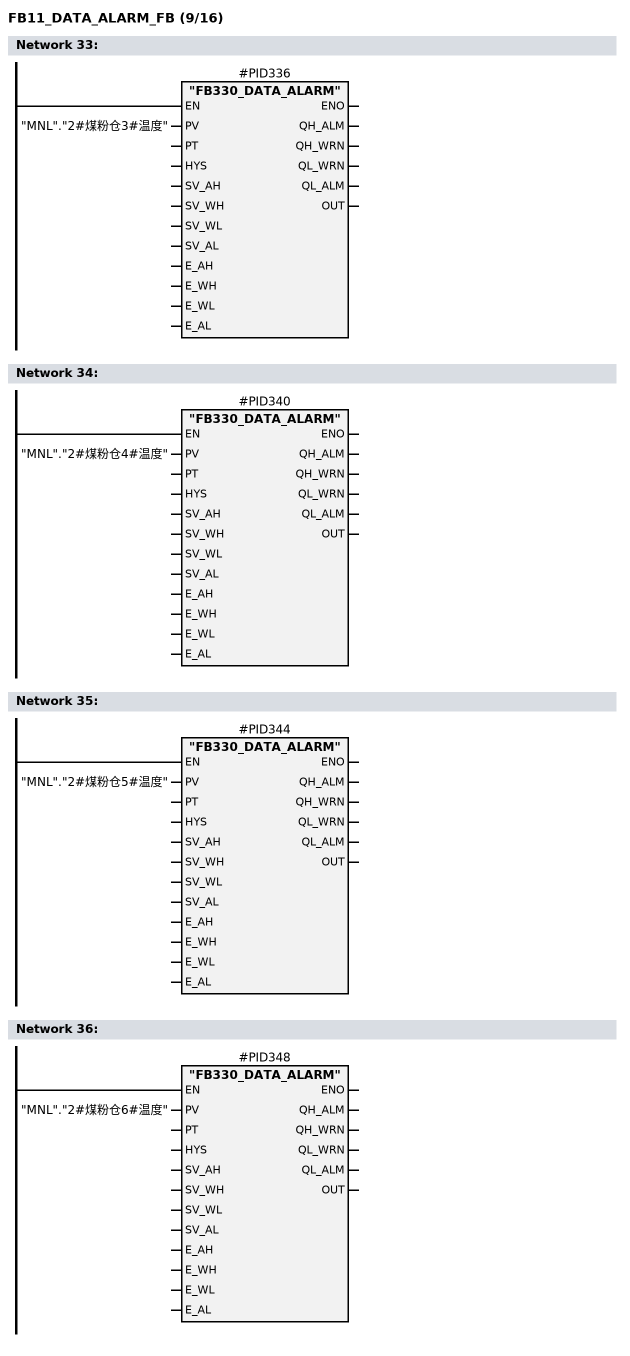
   RUNG wire#powerrail
      #PID336(PV := "MNL"."2#煤粉仓3#温度", PT :=, HYS :=, SV_AH :=, SV_WH :=, SV_WL :=, SV_AL :=, E_AH :=, E_WH :=, E_WL :=, E_AL :=, QH_ALM =>, QH_WRN =>, QL_WRN =>, QL_ALM =>, OUT =>)
   END_RUNG
   // the same network as SCL:
   #PID336(PV := "MNL"."2#煤粉仓3#温度");   // "FB330_DATA_ALARM"
END_REGION

REGION Network 34
   RUNG wire#powerrail
      #PID340(PV := "MNL"."2#煤粉仓4#温度", PT :=, HYS :=, SV_AH :=, SV_WH :=, SV_WL :=, SV_AL :=, E_AH :=, E_WH :=, E_WL :=, E_AL :=, QH_ALM =>, QH_WRN =>, QL_WRN =>, QL_ALM =>, OUT =>)
   END_RUNG
   // the same network as SCL:
   #PID340(PV := "MNL"."2#煤粉仓4#温度");   // "FB330_DATA_ALARM"
END_REGION

REGION Network 35
   RUNG wire#powerrail
      #PID344(PV := "MNL"."2#煤粉仓5#温度", PT :=, HYS :=, SV_AH :=, SV_WH :=, SV_WL :=, SV_AL :=, E_AH :=, E_WH :=, E_WL :=, E_AL :=, QH_ALM =>, QH_WRN =>, QL_WRN =>, QL_ALM =>, OUT =>)
   END_RUNG
   // the same network as SCL:
   #PID344(PV := "MNL"."2#煤粉仓5#温度");   // "FB330_DATA_ALARM"
END_REGION

REGION Network 36
   RUNG wire#powerrail
      #PID348(PV := "MNL"."2#煤粉仓6#温度", PT :=, HYS :=, SV_AH :=, SV_WH :=, SV_WL :=, SV_AL :=, E_AH :=, E_WH :=, E_WL :=, E_AL :=, QH_ALM =>, QH_WRN =>, QL_WRN =>, QL_ALM =>, OUT =>)
   END_RUNG
   // the same network as SCL:
   #PID348(PV := "MNL"."2#煤粉仓6#温度");   // "FB330_DATA_ALARM"
END_REGION

REGION Network 37
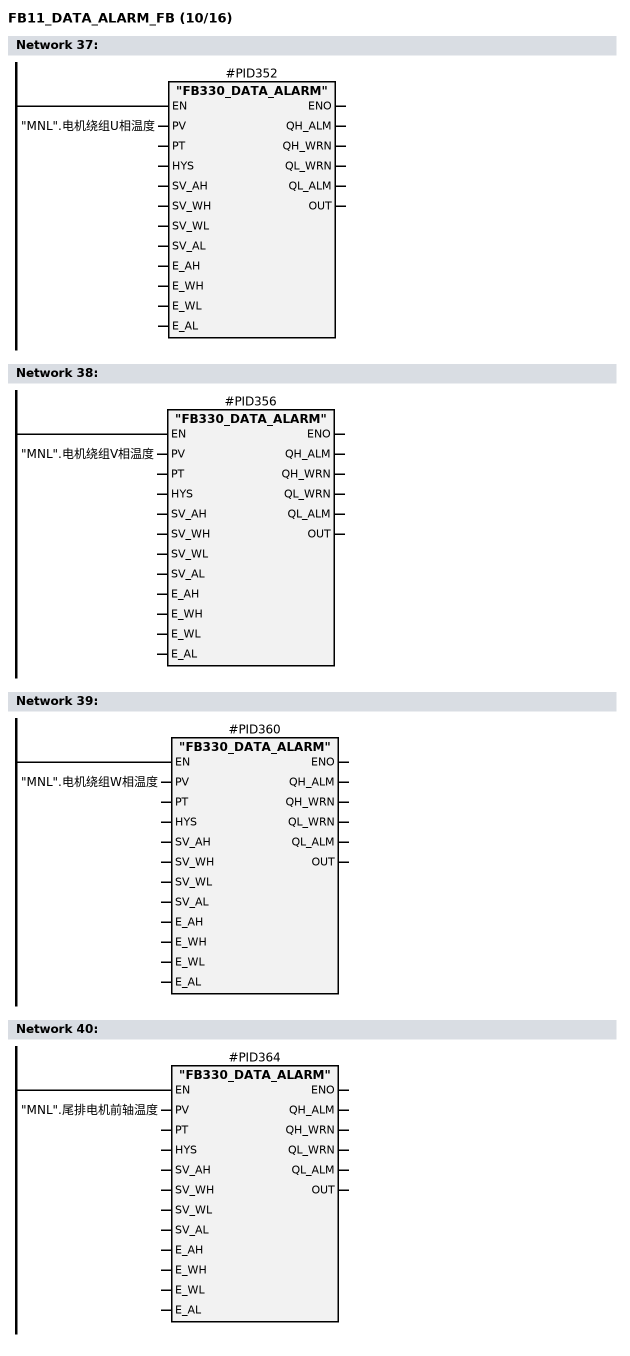
   RUNG wire#powerrail
      #PID352(PV := "MNL".电机绕组U相温度, PT :=, HYS :=, SV_AH :=, SV_WH :=, SV_WL :=, SV_AL :=, E_AH :=, E_WH :=, E_WL :=, E_AL :=, QH_ALM =>, QH_WRN =>, QL_WRN =>, QL_ALM =>, OUT =>)
   END_RUNG
   // the same network as SCL:
   #PID352(PV := "MNL".电机绕组U相温度);   // "FB330_DATA_ALARM"
END_REGION

REGION Network 38
   RUNG wire#powerrail
      #PID356(PV := "MNL".电机绕组V相温度, PT :=, HYS :=, SV_AH :=, SV_WH :=, SV_WL :=, SV_AL :=, E_AH :=, E_WH :=, E_WL :=, E_AL :=, QH_ALM =>, QH_WRN =>, QL_WRN =>, QL_ALM =>, OUT =>)
   END_RUNG
   // the same network as SCL:
   #PID356(PV := "MNL".电机绕组V相温度);   // "FB330_DATA_ALARM"
END_REGION

REGION Network 39
   RUNG wire#powerrail
      #PID360(PV := "MNL".电机绕组W相温度, PT :=, HYS :=, SV_AH :=, SV_WH :=, SV_WL :=, SV_AL :=, E_AH :=, E_WH :=, E_WL :=, E_AL :=, QH_ALM =>, QH_WRN =>, QL_WRN =>, QL_ALM =>, OUT =>)
   END_RUNG
   // the same network as SCL:
   #PID360(PV := "MNL".电机绕组W相温度);   // "FB330_DATA_ALARM"
END_REGION

REGION Network 40
   RUNG wire#powerrail
      #PID364(PV := "MNL".尾排电机前轴温度, PT :=, HYS :=, SV_AH :=, SV_WH :=, SV_WL :=, SV_AL :=, E_AH :=, E_WH :=, E_WL :=, E_AL :=, QH_ALM =>, QH_WRN =>, QL_WRN =>, QL_ALM =>, OUT =>)
   END_RUNG
   // the same network as SCL:
   #PID364(PV := "MNL".尾排电机前轴温度);   // "FB330_DATA_ALARM"
END_REGION

REGION Network 41
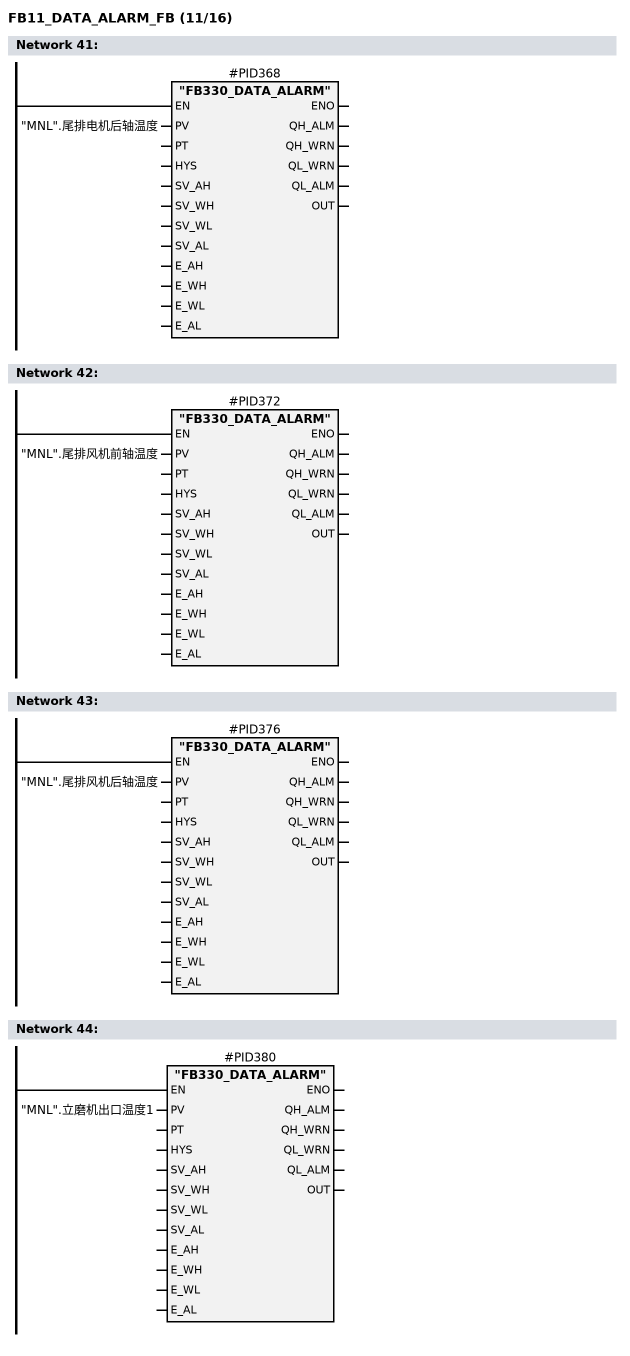
   RUNG wire#powerrail
      #PID368(PV := "MNL".尾排电机后轴温度, PT :=, HYS :=, SV_AH :=, SV_WH :=, SV_WL :=, SV_AL :=, E_AH :=, E_WH :=, E_WL :=, E_AL :=, QH_ALM =>, QH_WRN =>, QL_WRN =>, QL_ALM =>, OUT =>)
   END_RUNG
   // the same network as SCL:
   #PID368(PV := "MNL".尾排电机后轴温度);   // "FB330_DATA_ALARM"
END_REGION

REGION Network 42
   RUNG wire#powerrail
      #PID372(PV := "MNL".尾排风机前轴温度, PT :=, HYS :=, SV_AH :=, SV_WH :=, SV_WL :=, SV_AL :=, E_AH :=, E_WH :=, E_WL :=, E_AL :=, QH_ALM =>, QH_WRN =>, QL_WRN =>, QL_ALM =>, OUT =>)
   END_RUNG
   // the same network as SCL:
   #PID372(PV := "MNL".尾排风机前轴温度);   // "FB330_DATA_ALARM"
END_REGION

REGION Network 43
   RUNG wire#powerrail
      #PID376(PV := "MNL".尾排风机后轴温度, PT :=, HYS :=, SV_AH :=, SV_WH :=, SV_WL :=, SV_AL :=, E_AH :=, E_WH :=, E_WL :=, E_AL :=, QH_ALM =>, QH_WRN =>, QL_WRN =>, QL_ALM =>, OUT =>)
   END_RUNG
   // the same network as SCL:
   #PID376(PV := "MNL".尾排风机后轴温度);   // "FB330_DATA_ALARM"
END_REGION

REGION Network 44
   RUNG wire#powerrail
      #PID380(PV := "MNL".立磨机出口温度1, PT :=, HYS :=, SV_AH :=, SV_WH :=, SV_WL :=, SV_AL :=, E_AH :=, E_WH :=, E_WL :=, E_AL :=, QH_ALM =>, QH_WRN =>, QL_WRN =>, QL_ALM =>, OUT =>)
   END_RUNG
   // the same network as SCL:
   #PID380(PV := "MNL".立磨机出口温度1);   // "FB330_DATA_ALARM"
END_REGION

REGION Network 45
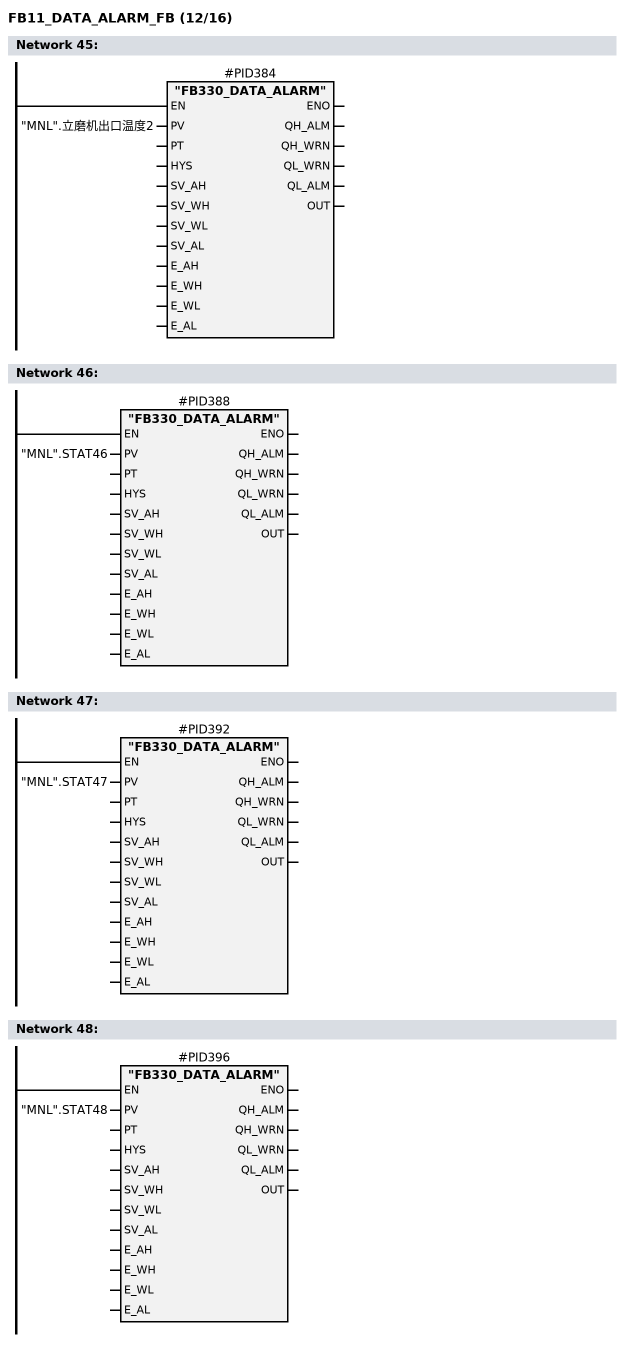
   RUNG wire#powerrail
      #PID384(PV := "MNL".立磨机出口温度2, PT :=, HYS :=, SV_AH :=, SV_WH :=, SV_WL :=, SV_AL :=, E_AH :=, E_WH :=, E_WL :=, E_AL :=, QH_ALM =>, QH_WRN =>, QL_WRN =>, QL_ALM =>, OUT =>)
   END_RUNG
   // the same network as SCL:
   #PID384(PV := "MNL".立磨机出口温度2);   // "FB330_DATA_ALARM"
END_REGION

REGION Network 46
   RUNG wire#powerrail
      #PID388(PV := "MNL".STAT46, PT :=, HYS :=, SV_AH :=, SV_WH :=, SV_WL :=, SV_AL :=, E_AH :=, E_WH :=, E_WL :=, E_AL :=, QH_ALM =>, QH_WRN =>, QL_WRN =>, QL_ALM =>, OUT =>)
   END_RUNG
   // the same network as SCL:
   #PID388(PV := "MNL".STAT46);   // "FB330_DATA_ALARM"
END_REGION

REGION Network 47
   RUNG wire#powerrail
      #PID392(PV := "MNL".STAT47, PT :=, HYS :=, SV_AH :=, SV_WH :=, SV_WL :=, SV_AL :=, E_AH :=, E_WH :=, E_WL :=, E_AL :=, QH_ALM =>, QH_WRN =>, QL_WRN =>, QL_ALM =>, OUT =>)
   END_RUNG
   // the same network as SCL:
   #PID392(PV := "MNL".STAT47);   // "FB330_DATA_ALARM"
END_REGION

REGION Network 48
   RUNG wire#powerrail
      #PID396(PV := "MNL".STAT48, PT :=, HYS :=, SV_AH :=, SV_WH :=, SV_WL :=, SV_AL :=, E_AH :=, E_WH :=, E_WL :=, E_AL :=, QH_ALM =>, QH_WRN =>, QL_WRN =>, QL_ALM =>, OUT =>)
   END_RUNG
   // the same network as SCL:
   #PID396(PV := "MNL".STAT48);   // "FB330_DATA_ALARM"
END_REGION

REGION Network 49
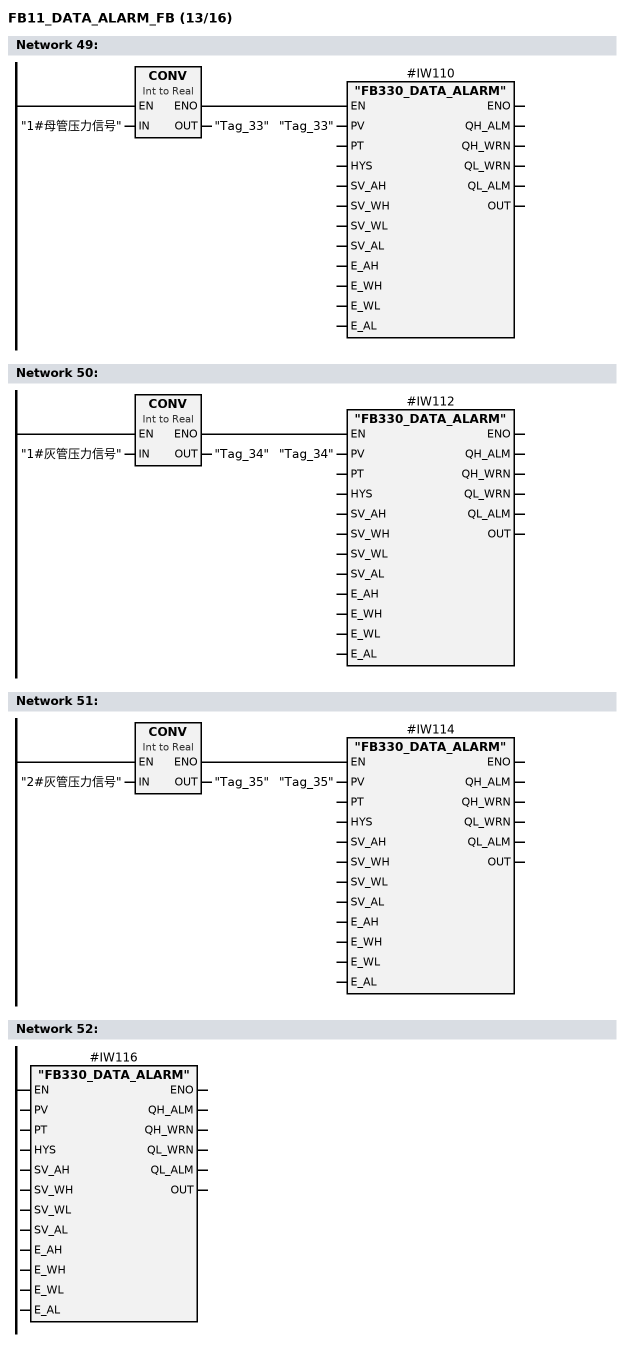
   RUNG wire#powerrail
      { S7_Templates := "[SrcType := Int, DestType := Real]" } Convert(in := "1#母管压力信号", out => "Tag_33")
      #IW110(PV := "Tag_33", PT :=, HYS :=, SV_AH :=, SV_WH :=, SV_WL :=, SV_AL :=, E_AH :=, E_WH :=, E_WL :=, E_AL :=, QH_ALM =>, QH_WRN =>, QL_WRN =>, QL_ALM =>, OUT =>)
   END_RUNG
   // the same network as SCL:
   "Tag_33" := INT_TO_REAL("1#母管压力信号");
   #IW110(PV := "Tag_33");   // "FB330_DATA_ALARM"
END_REGION

REGION Network 50
   RUNG wire#powerrail
      { S7_Templates := "[SrcType := Int, DestType := Real]" } Convert(in := "1#灰管压力信号", out => "Tag_34")
      #IW112(PV := "Tag_34", PT :=, HYS :=, SV_AH :=, SV_WH :=, SV_WL :=, SV_AL :=, E_AH :=, E_WH :=, E_WL :=, E_AL :=, QH_ALM =>, QH_WRN =>, QL_WRN =>, QL_ALM =>, OUT =>)
   END_RUNG
   // the same network as SCL:
   "Tag_34" := INT_TO_REAL("1#灰管压力信号");
   #IW112(PV := "Tag_34");   // "FB330_DATA_ALARM"
END_REGION

REGION Network 51
   RUNG wire#powerrail
      { S7_Templates := "[SrcType := Int, DestType := Real]" } Convert(in := "2#灰管压力信号", out => "Tag_35")
      #IW114(PV := "Tag_35", PT :=, HYS :=, SV_AH :=, SV_WH :=, SV_WL :=, SV_AL :=, E_AH :=, E_WH :=, E_WL :=, E_AL :=, QH_ALM =>, QH_WRN =>, QL_WRN =>, QL_ALM =>, OUT =>)
   END_RUNG
   // the same network as SCL:
   "Tag_35" := INT_TO_REAL("2#灰管压力信号");
   #IW114(PV := "Tag_35");   // "FB330_DATA_ALARM"
END_REGION

REGION Network 52
   RUNG wire#powerrail
      #IW116(PV :=, PT :=, HYS :=, SV_AH :=, SV_WH :=, SV_WL :=, SV_AL :=, E_AH :=, E_WH :=, E_WL :=, E_AL :=, QH_ALM =>, QH_WRN =>, QL_WRN =>, QL_ALM =>, OUT =>)
   END_RUNG
   // the same network as SCL:
   #IW116();   // "FB330_DATA_ALARM"
END_REGION

REGION Network 53
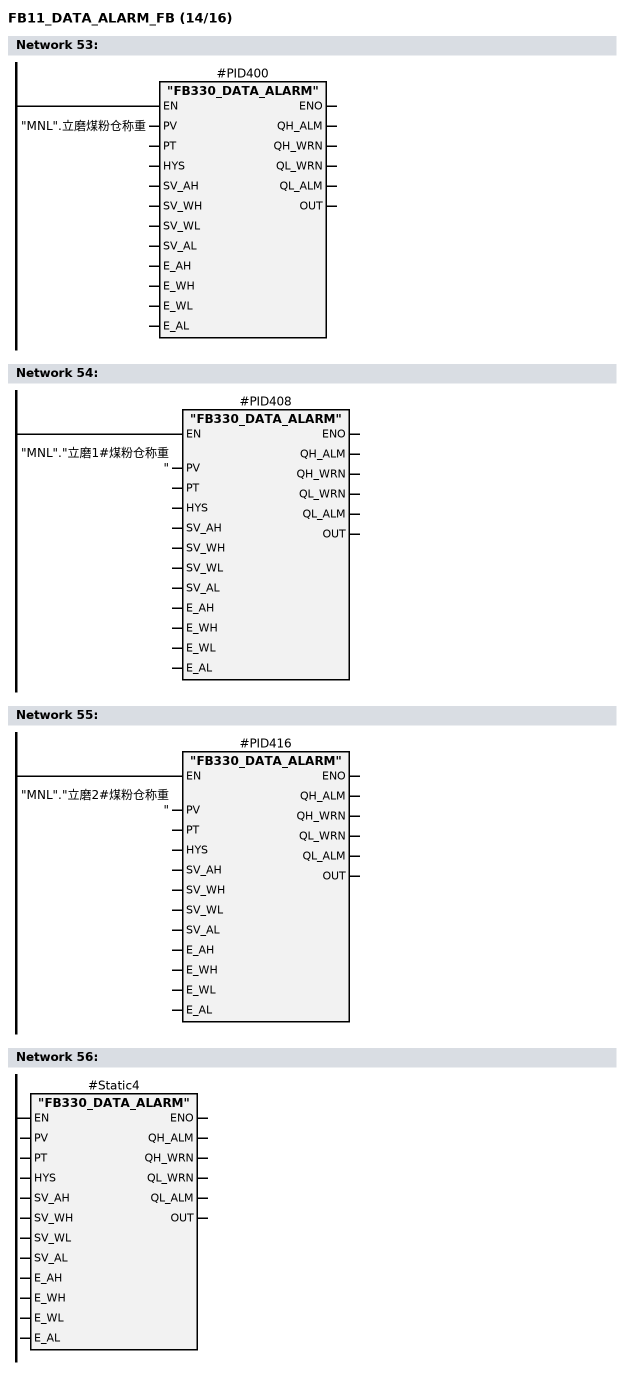
   RUNG wire#powerrail
      #PID400(PV := "MNL".立磨煤粉仓称重, PT :=, HYS :=, SV_AH :=, SV_WH :=, SV_WL :=, SV_AL :=, E_AH :=, E_WH :=, E_WL :=, E_AL :=, QH_ALM =>, QH_WRN =>, QL_WRN =>, QL_ALM =>, OUT =>)
   END_RUNG
   // the same network as SCL:
   #PID400(PV := "MNL".立磨煤粉仓称重);   // "FB330_DATA_ALARM"
END_REGION

REGION Network 54
   RUNG wire#powerrail
      #PID408(PV := "MNL"."立磨1#煤粉仓称重", PT :=, HYS :=, SV_AH :=, SV_WH :=, SV_WL :=, SV_AL :=, E_AH :=, E_WH :=, E_WL :=, E_AL :=, QH_ALM =>, QH_WRN =>, QL_WRN =>, QL_ALM =>, OUT =>)
   END_RUNG
   // the same network as SCL:
   #PID408(PV := "MNL"."立磨1#煤粉仓称重");   // "FB330_DATA_ALARM"
END_REGION

REGION Network 55
   RUNG wire#powerrail
      #PID416(PV := "MNL"."立磨2#煤粉仓称重", PT :=, HYS :=, SV_AH :=, SV_WH :=, SV_WL :=, SV_AL :=, E_AH :=, E_WH :=, E_WL :=, E_AL :=, QH_ALM =>, QH_WRN =>, QL_WRN =>, QL_ALM =>, OUT =>)
   END_RUNG
   // the same network as SCL:
   #PID416(PV := "MNL"."立磨2#煤粉仓称重");   // "FB330_DATA_ALARM"
END_REGION

REGION Network 56
   RUNG wire#powerrail
      #Static4(PV :=, PT :=, HYS :=, SV_AH :=, SV_WH :=, SV_WL :=, SV_AL :=, E_AH :=, E_WH :=, E_WL :=, E_AL :=, QH_ALM =>, QH_WRN =>, QL_WRN =>, QL_ALM =>, OUT =>)
   END_RUNG
   // the same network as SCL:
   #Static4();   // "FB330_DATA_ALARM"
END_REGION

REGION Network 57
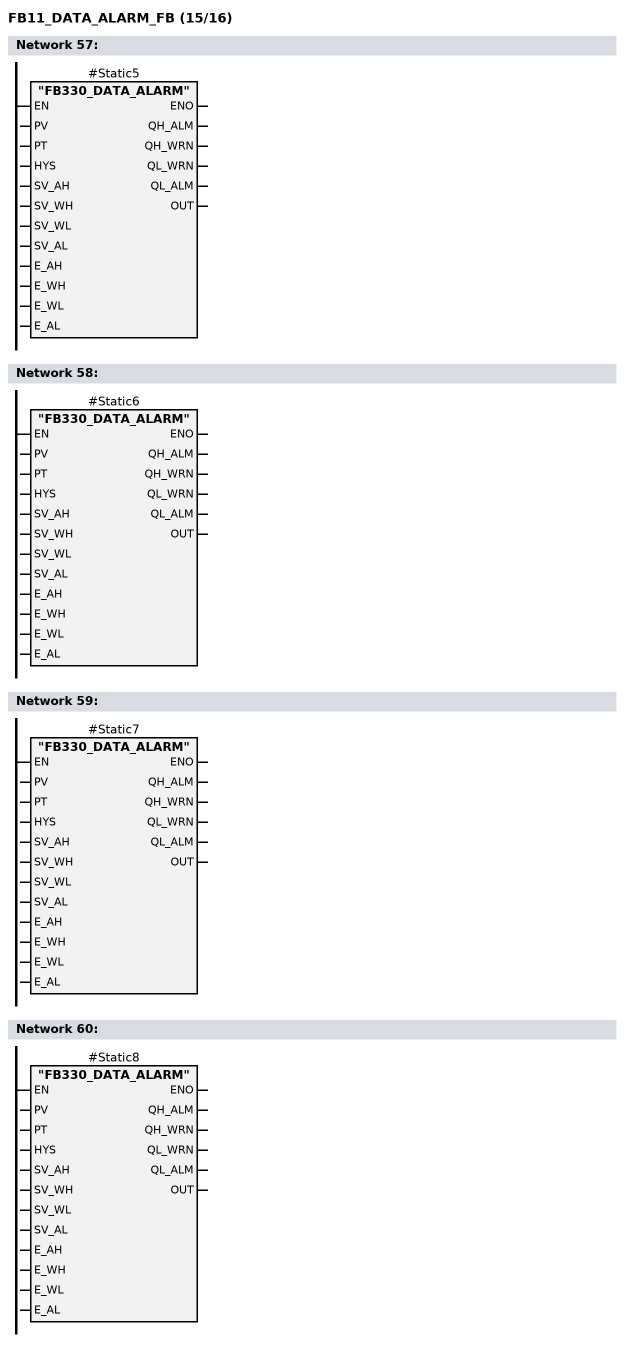
   RUNG wire#powerrail
      #Static5(PV :=, PT :=, HYS :=, SV_AH :=, SV_WH :=, SV_WL :=, SV_AL :=, E_AH :=, E_WH :=, E_WL :=, E_AL :=, QH_ALM =>, QH_WRN =>, QL_WRN =>, QL_ALM =>, OUT =>)
   END_RUNG
   // the same network as SCL:
   #Static5();   // "FB330_DATA_ALARM"
END_REGION

REGION Network 58
   RUNG wire#powerrail
      #Static6(PV :=, PT :=, HYS :=, SV_AH :=, SV_WH :=, SV_WL :=, SV_AL :=, E_AH :=, E_WH :=, E_WL :=, E_AL :=, QH_ALM =>, QH_WRN =>, QL_WRN =>, QL_ALM =>, OUT =>)
   END_RUNG
   // the same network as SCL:
   #Static6();   // "FB330_DATA_ALARM"
END_REGION

REGION Network 59
   RUNG wire#powerrail
      #Static7(PV :=, PT :=, HYS :=, SV_AH :=, SV_WH :=, SV_WL :=, SV_AL :=, E_AH :=, E_WH :=, E_WL :=, E_AL :=, QH_ALM =>, QH_WRN =>, QL_WRN =>, QL_ALM =>, OUT =>)
   END_RUNG
   // the same network as SCL:
   #Static7();   // "FB330_DATA_ALARM"
END_REGION

REGION Network 60
   RUNG wire#powerrail
      #Static8(PV :=, PT :=, HYS :=, SV_AH :=, SV_WH :=, SV_WL :=, SV_AL :=, E_AH :=, E_WH :=, E_WL :=, E_AL :=, QH_ALM =>, QH_WRN =>, QL_WRN =>, QL_ALM =>, OUT =>)
   END_RUNG
   // the same network as SCL:
   #Static8();   // "FB330_DATA_ALARM"
END_REGION

REGION Network 61
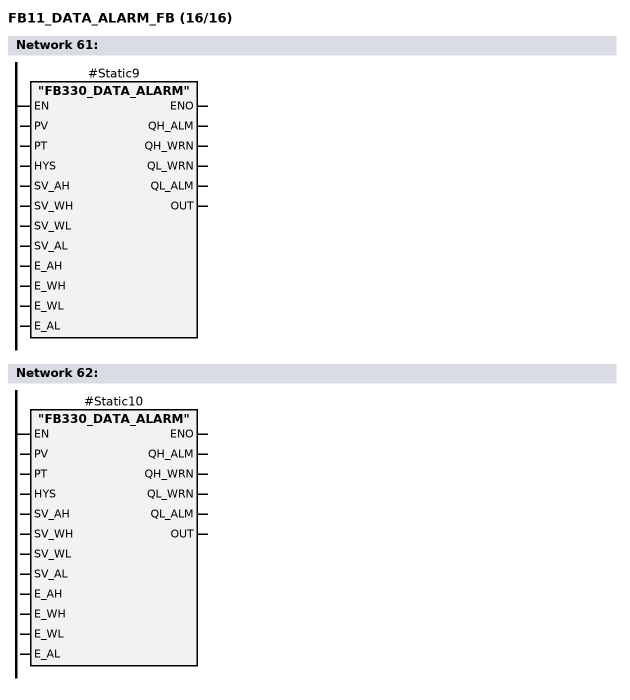
   RUNG wire#powerrail
      #Static9(PV :=, PT :=, HYS :=, SV_AH :=, SV_WH :=, SV_WL :=, SV_AL :=, E_AH :=, E_WH :=, E_WL :=, E_AL :=, QH_ALM =>, QH_WRN =>, QL_WRN =>, QL_ALM =>, OUT =>)
   END_RUNG
   // the same network as SCL:
   #Static9();   // "FB330_DATA_ALARM"
END_REGION

REGION Network 62
   RUNG wire#powerrail
      #Static10(PV :=, PT :=, HYS :=, SV_AH :=, SV_WH :=, SV_WL :=, SV_AL :=, E_AH :=, E_WH :=, E_WL :=, E_AL :=, QH_ALM =>, QH_WRN =>, QL_WRN =>, QL_ALM =>, OUT =>)
   END_RUNG
   // the same network as SCL:
   #Static10();   // "FB330_DATA_ALARM"
END_REGION
END_FUNCTION_BLOCK

FUNCTION_BLOCK "阀门控制块"   // FB300, LAD
{ S7_Optimized_Access := 'TRUE' }
VERSION : 0.1
   VAR_INPUT
      LR : Bool;
      V_OPEN : Bool;
      V_CLOSE : Bool;
      HMI_OPEN : Bool;
      HMI_CLOSE : Bool;
   END_VAR
   VAR_OUTPUT
      OUT_OP_PULSE : Bool;
      OUT_CL_PULSE : Bool;
   END_VAR
   VAR_IN_OUT
      OUT_HOLD : Bool;
   END_VAR
BEGIN

REGION Network 1
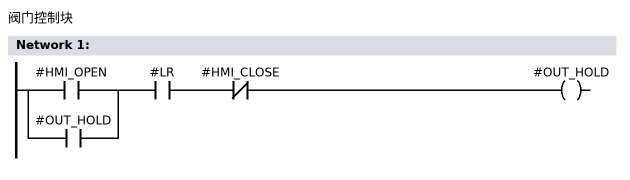
   RUNG wire#powerrail
      Contact( #HMI_OPEN )
      wire#w1
      Contact( #LR )
      I_Contact( #HMI_CLOSE )
      Coil( #OUT_HOLD )
   END_RUNG
   RUNG wire#powerrail
      Contact( #OUT_HOLD )
   END_RUNG wire#w1
   // the same network as SCL:
   #OUT_HOLD := (#HMI_OPEN OR #OUT_HOLD) AND #LR AND NOT #HMI_CLOSE;
END_REGION
END_FUNCTION_BLOCK

FUNCTION_BLOCK "FB330_DATA_ALARM"   // FB330, LAD
{ S7_Optimized_Access := 'FALSE' }
VERSION : 0.1
// REAL的报警块
   VAR_INPUT
      PV : Real;   // 过程值
      PT : Real := 1.0;   // 系数
      HYS : Real;   // 回差值
      SV_AH : Real;   // 高报警设定值
      SV_WH : Real;   // 高警告设定值
      SV_WL : Real;   // 低警告设定值
      SV_AL : Real;   // 低报警设定值
      E_AH : Bool;   // 高报警使能
      E_WH : Bool;   // 高警告使能
      E_WL : Bool;   // 低警告使能
      E_AL : Bool;   // 低报警使能
   END_VAR
   VAR_OUTPUT
      QH_ALM : Bool;   // 高报警输出
      QH_WRN : Bool;   // 高警告输出
      QL_WRN : Bool;   // 低警告输出
      QL_ALM : Bool;   // 低报警输出
      OUT : Real;   // 输出
   END_VAR
   VAR
      SR1 : Bool;
      SR2 : Bool;
      SR3 : Bool;
      SR4 : Bool;
   END_VAR
   VAR_TEMP
      TEMP_AH : Real;
      TEMP_WH : Real;
      TEMP_AL : Real;
      TEMP_WL : Real;
      TEMP_OUT : Real;
   END_VAR
BEGIN

REGION Network 1
   // 系数转换
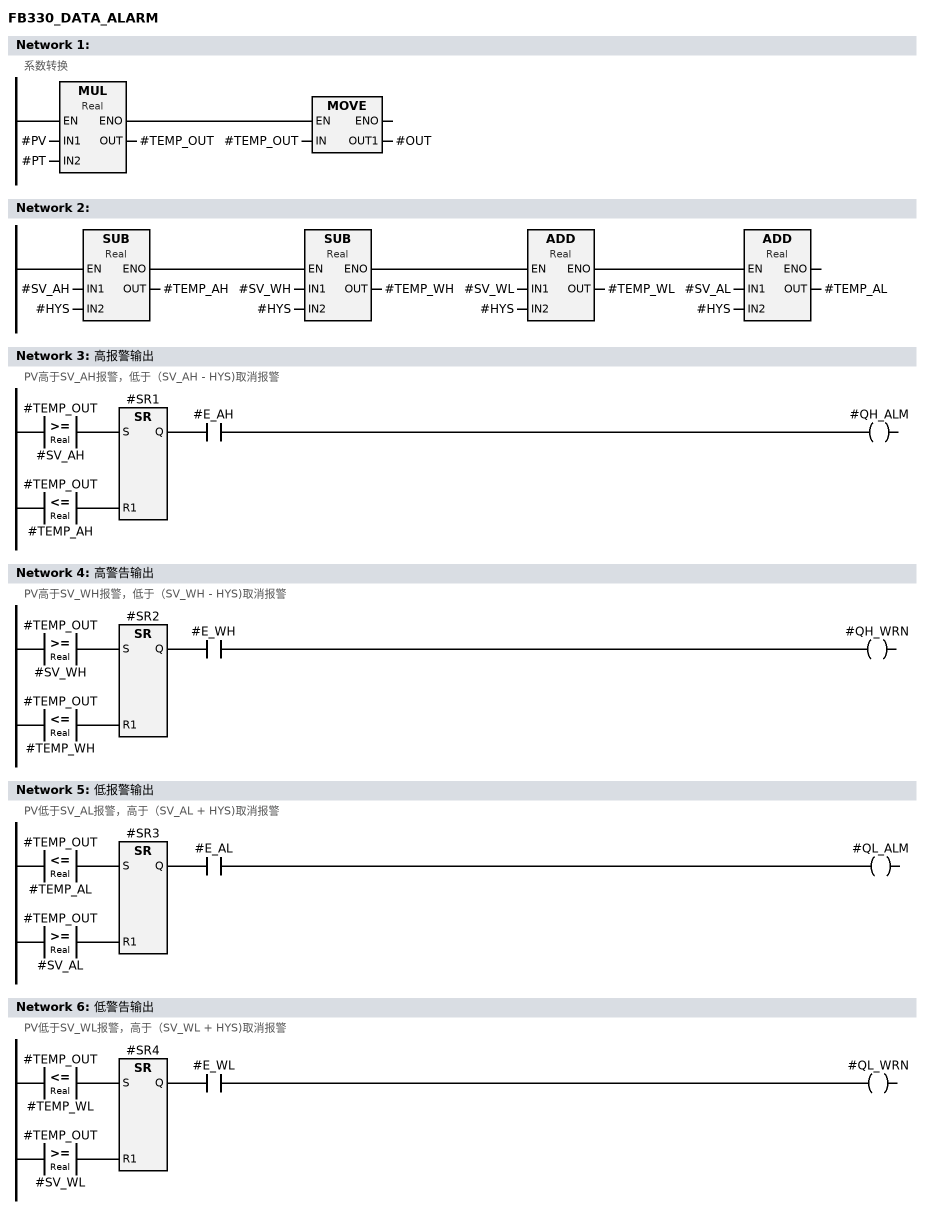
   RUNG wire#powerrail
      { S7_Templates := "SrcType := Real"; S7_GenerateENO := "TRUE" } Mul(in1 := #PV, in2 := #PT, out => #TEMP_OUT)
      { S7_GenerateENO := "TRUE" } Move(in := #TEMP_OUT, out1 => #OUT)
   END_RUNG
   // the same network as SCL:
   // ENO of a box is taken as its EN; it also drops when the box reports an error
   #TEMP_OUT := #PV * #PT;
   #OUT := #TEMP_OUT;
END_REGION

REGION Network 2
   RUNG wire#powerrail
      { S7_Templates := "SrcType := Real"; S7_GenerateENO := "TRUE" } Sub(in1 := #SV_AH, in2 := #HYS, out => #TEMP_AH)
      { S7_Templates := "SrcType := Real"; S7_GenerateENO := "TRUE" } Sub(in1 := #SV_WH, in2 := #HYS, out => #TEMP_WH)
      { S7_Templates := "SrcType := Real"; S7_GenerateENO := "TRUE" } Add(in1 := #SV_WL, in2 := #HYS, out => #TEMP_WL)
      { S7_Templates := "SrcType := Real"; S7_GenerateENO := "TRUE" } Add(in1 := #SV_AL, in2 := #HYS, out => #TEMP_AL)
   END_RUNG
   // the same network as SCL:
   // ENO of a box is taken as its EN; it also drops when the box reports an error
   #TEMP_AH := #SV_AH - #HYS;
   #TEMP_WH := #SV_WH - #HYS;
   #TEMP_WL := #SV_WL + #HYS;
   #TEMP_AL := #SV_AL + #HYS;
END_REGION

REGION Network 3: 高报警输出
   // PV高于SV_AH报警，低于（SV_AH - HYS)取消报警
   RUNG wire#powerrail
      { S7_Templates := "SrcType := Real" } GE_Contact(in1 := #TEMP_OUT, in2 := #SV_AH)
      S_SR(operand := #SR1, r1 := wire#w1)
      Contact( #E_AH )
      Coil( #QH_ALM )
   END_RUNG
   RUNG wire#powerrail
      { S7_Templates := "SrcType := Real" } LE_Contact(in1 := #TEMP_OUT, in2 := #TEMP_AH)
   END_RUNG wire#w1
   // the same network as SCL:
   IF #TEMP_OUT >= #SV_AH THEN
       #SR1 := TRUE;   // SR flip-flop
   END_IF;
   IF #TEMP_OUT <= #TEMP_AH THEN #SR1 := FALSE; END_IF;
   #QH_ALM := #SR1 AND #E_AH;
END_REGION

REGION Network 4: 高警告输出
   // PV高于SV_WH报警，低于（SV_WH - HYS)取消报警
   RUNG wire#powerrail
      { S7_Templates := "SrcType := Real" } GE_Contact(in1 := #TEMP_OUT, in2 := #SV_WH)
      S_SR(operand := #SR2, r1 := wire#w1)
      Contact( #E_WH )
      Coil( #QH_WRN )
   END_RUNG
   RUNG wire#powerrail
      { S7_Templates := "SrcType := Real" } LE_Contact(in1 := #TEMP_OUT, in2 := #TEMP_WH)
   END_RUNG wire#w1
   // the same network as SCL:
   IF #TEMP_OUT >= #SV_WH THEN
       #SR2 := TRUE;   // SR flip-flop
   END_IF;
   IF #TEMP_OUT <= #TEMP_WH THEN #SR2 := FALSE; END_IF;
   #QH_WRN := #SR2 AND #E_WH;
END_REGION

REGION Network 5: 低报警输出
   // PV低于SV_AL报警，高于（SV_AL + HYS)取消报警
   RUNG wire#powerrail
      { S7_Templates := "SrcType := Real" } LE_Contact(in1 := #TEMP_OUT, in2 := #TEMP_AL)
      S_SR(operand := #SR3, r1 := wire#w1)
      Contact( #E_AL )
      Coil( #QL_ALM )
   END_RUNG
   RUNG wire#powerrail
      { S7_Templates := "SrcType := Real" } GE_Contact(in1 := #TEMP_OUT, in2 := #SV_AL)
   END_RUNG wire#w1
   // the same network as SCL:
   IF #TEMP_OUT <= #TEMP_AL THEN
       #SR3 := TRUE;   // SR flip-flop
   END_IF;
   IF #TEMP_OUT >= #SV_AL THEN #SR3 := FALSE; END_IF;
   #QL_ALM := #SR3 AND #E_AL;
END_REGION

REGION Network 6: 低警告输出
   // PV低于SV_WL报警，高于（SV_WL + HYS)取消报警
   RUNG wire#powerrail
      { S7_Templates := "SrcType := Real" } LE_Contact(in1 := #TEMP_OUT, in2 := #TEMP_WL)
      S_SR(operand := #SR4, r1 := wire#w1)
      Contact( #E_WL )
      Coil( #QL_WRN )
   END_RUNG
   RUNG wire#powerrail
      { S7_Templates := "SrcType := Real" } GE_Contact(in1 := #TEMP_OUT, in2 := #SV_WL)
   END_RUNG wire#w1
   // the same network as SCL:
   IF #TEMP_OUT <= #TEMP_WL THEN
       #SR4 := TRUE;   // SR flip-flop
   END_IF;
   IF #TEMP_OUT >= #SV_WL THEN #SR4 := FALSE; END_IF;
   #QL_WRN := #SR4 AND #E_WL;
END_REGION
END_FUNCTION_BLOCK

FUNCTION "电机控制" : Void   // FC1, LAD
{ S7_Optimized_Access := 'FALSE' }
VERSION : 0.1
   VAR_TEMP   // added for the SCL form of the ladder/FBD networks
      _w1 : Bool;
      _s5time1 : S5Time;
      _w2 : Bool;
   END_VAR
BEGIN

REGION Network 2
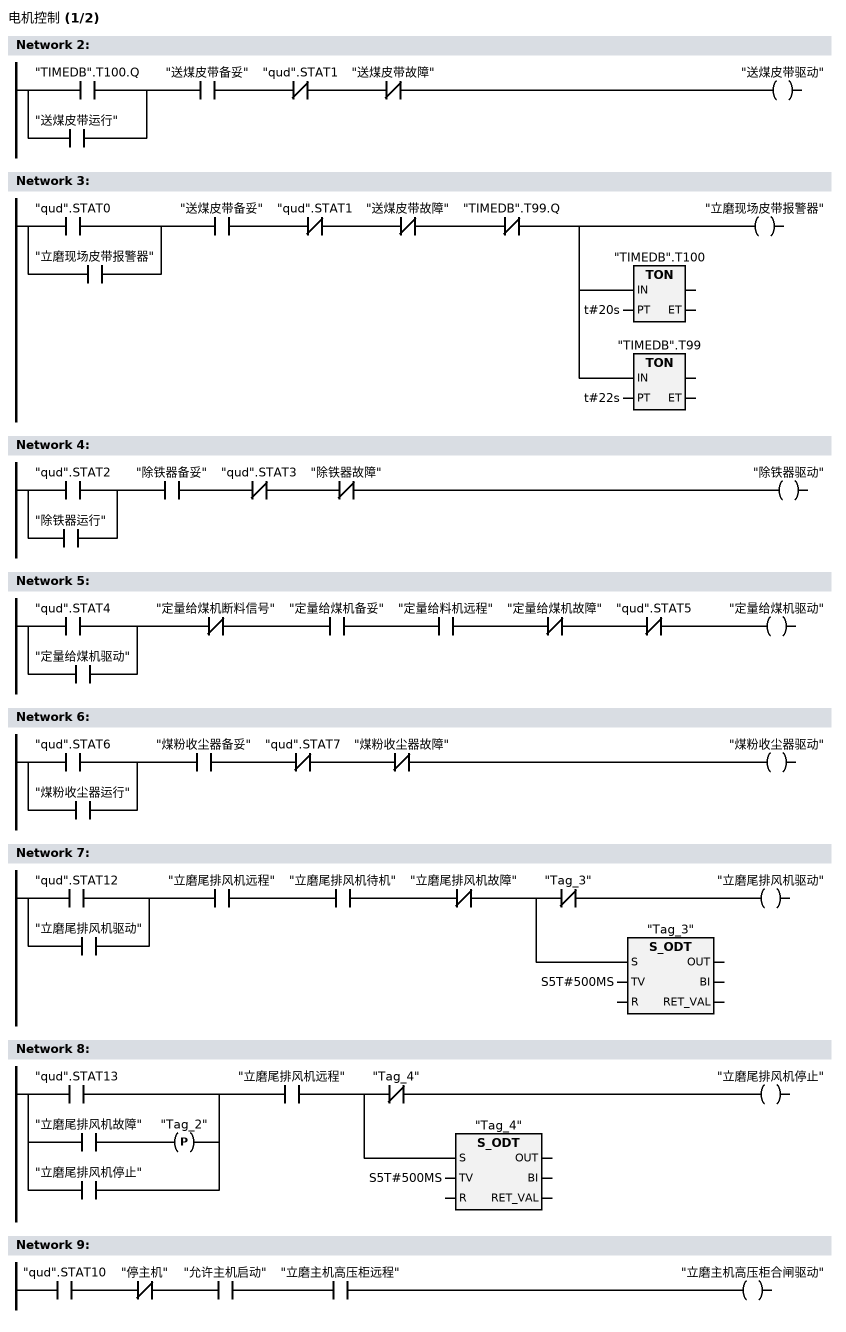
   RUNG wire#powerrail
      Contact( "TIMEDB".T100.Q )
      wire#w1
      Contact( "送煤皮带备妥" )
      I_Contact( "qud".STAT1 )
      I_Contact( "送煤皮带故障" )
      Coil( "送煤皮带驱动" )
   END_RUNG
   RUNG wire#powerrail
      Contact( "送煤皮带运行" )
   END_RUNG wire#w1
   // the same network as SCL:
   "送煤皮带驱动" := ("TIMEDB".T100.Q OR "送煤皮带运行") AND "送煤皮带备妥" AND NOT "qud".STAT1 AND NOT "送煤皮带故障";
END_REGION

REGION Network 3
   "立磨现场皮带报警器" := ("qud".STAT0 OR "立磨现场皮带报警器") AND "送煤皮带备妥" AND NOT "qud".STAT1 AND NOT "送煤皮带故障" AND NOT "TIMEDB".T99.Q;
   "TIMEDB".T100.TON(IN := "立磨现场皮带报警器", PT := t#20s);
   "TIMEDB".T99.TON(IN := "立磨现场皮带报警器", PT := t#22s);
END_REGION

REGION Network 4
   RUNG wire#powerrail
      Contact( "qud".STAT2 )
      wire#w1
      Contact( "除铁器备妥" )
      I_Contact( "qud".STAT3 )
      I_Contact( "除铁器故障" )
      Coil( "除铁器驱动" )
   END_RUNG
   RUNG wire#powerrail
      Contact( "除铁器运行" )
   END_RUNG wire#w1
   // the same network as SCL:
   "除铁器驱动" := ("qud".STAT2 OR "除铁器运行") AND "除铁器备妥" AND NOT "qud".STAT3 AND NOT "除铁器故障";
END_REGION

REGION Network 5
   RUNG wire#powerrail
      Contact( "qud".STAT4 )
      wire#w1
      I_Contact( "定量给煤机断料信号" )
      Contact( "定量给煤机备妥" )
      Contact( "定量给料机远程" )
      I_Contact( "定量给煤机故障" )
      I_Contact( "qud".STAT5 )
      Coil( "定量给煤机驱动" )
   END_RUNG
   RUNG wire#powerrail
      Contact( "定量给煤机驱动" )
   END_RUNG wire#w1
   // the same network as SCL:
   "定量给煤机驱动" := ("qud".STAT4 OR "定量给煤机驱动") AND NOT "定量给煤机断料信号" AND "定量给煤机备妥" AND "定量给料机远程" AND NOT "定量给煤机故障" AND NOT "qud".STAT5;
END_REGION

REGION Network 6
   RUNG wire#powerrail
      Contact( "qud".STAT6 )
      wire#w1
      Contact( "煤粉收尘器备妥" )
      I_Contact( "qud".STAT7 )
      I_Contact( "煤粉收尘器故障" )
      Coil( "煤粉收尘器驱动" )
   END_RUNG
   RUNG wire#powerrail
      Contact( "煤粉收尘器运行" )
   END_RUNG wire#w1
   // the same network as SCL:
   "煤粉收尘器驱动" := ("qud".STAT6 OR "煤粉收尘器运行") AND "煤粉收尘器备妥" AND NOT "qud".STAT7 AND NOT "煤粉收尘器故障";
END_REGION

REGION Network 7
   RUNG wire#powerrail
      Contact( "qud".STAT12 )
      wire#w1
      Contact( "立磨尾排风机远程" )
      Contact( "立磨尾排风机待机" )
      I_Contact( "立磨尾排风机故障" )
      wire#w2
      I_Contact( "Tag_3" )
      Coil( "立磨尾排风机驱动" )
   END_RUNG
   RUNG wire#powerrail
      Contact( "立磨尾排风机驱动" )
   END_RUNG wire#w1
   RUNG wire#w2
      S_ODT(T_NO := "Tag_3", TV := S5T#500MS, R :=, BI =>, RET_VAL =>)
   END_RUNG
   // the same network as SCL:
   #_w1 := ("qud".STAT12 OR "立磨尾排风机驱动") AND "立磨尾排风机远程" AND "立磨尾排风机待机" AND NOT "立磨尾排风机故障";
   "立磨尾排风机驱动" := #_w1 AND NOT "Tag_3";
   #_s5time1 := S_ODT(T_NO := "Tag_3", TV := S5T#500MS, S := #_w1);
END_REGION

REGION Network 8
   RUNG wire#powerrail
      Contact( "qud".STAT13 )
      wire#w1
      Contact( "立磨尾排风机远程" )
      wire#w2
      I_Contact( "Tag_4" )
      Coil( "立磨尾排风机停止" )
   END_RUNG
   RUNG wire#powerrail
      Contact( "立磨尾排风机故障" )
      P_Trig( "Tag_2" )
   END_RUNG wire#w1
   RUNG wire#powerrail
      Contact( "立磨尾排风机停止" )
   END_RUNG wire#w1
   RUNG wire#w2
      S_ODT(T_NO := "Tag_4", TV := S5T#500MS, R :=, BI =>, RET_VAL =>)
   END_RUNG
   // the same network as SCL:
   #_w1 := "立磨尾排风机故障" AND NOT "Tag_2";   // rising edge
   "Tag_2" := "立磨尾排风机故障";
   #_w2 := ("qud".STAT13 OR #_w1 OR "立磨尾排风机停止") AND "立磨尾排风机远程";
   "立磨尾排风机停止" := #_w2 AND NOT "Tag_4";
   #_s5time1 := S_ODT(T_NO := "Tag_4", S := #_w2, TV := S5T#500MS);
END_REGION

REGION Network 9
   RUNG wire#powerrail
      Contact( "qud".STAT10 )
      I_Contact( "停主机" )
      Contact( "允许主机启动" )
      Contact( "立磨主机高压柜远程" )
      Coil( "立磨主机高压柜合闸驱动" )
   END_RUNG
   // the same network as SCL:
   "立磨主机高压柜合闸驱动" := "qud".STAT10 AND NOT "停主机" AND "允许主机启动" AND "立磨主机高压柜远程";
END_REGION

REGION Network 10
